      "1133_GTT_DETERMINE_EXCLUSIVITY"(TankID_InOperation := 11, DemandComplete := #GTT_OUT.GTT_DemandsCompleted[11], GTT_Exclusivity := #GTT_Exclusivity)
   END_RUNG
   RUNG wire#powerrail
      { S7_Templates := "SrcType := Int" } EQ_Contact(in1 := #GTT_Exclusivity.TankID_InOperation, in2 := 11)
   END_RUNG wire#w2
   RUNG wire#w2
      I_Coil( #DNC_5S_GTT.Reset )
   END_RUNG
   // the same network as SCL:
   #_w1 := (NOT #GTT_Exclusivity.Tank_Exclusivity AND #GTT_IN.GTT_Actuate[10] AND NOT #GTT_OUT.GTT_DemandsCompleted[10]) OR (#GTT_Exclusivity.TankID_InOperation = 10);
   #"5P_GTT_TimeSel" := "1135_VALVE_OPEN_CLOSE_TIME_SEL"(EN := #_w1,
                           ValveType := 0,
                           ValveDemand := #GTT_IN.GTT_ValveDemands[10],
                           OpenTime := "1096_ADJUSTABLE_CONSTANTS".BWTInletValveOpen_Time,
                           CloseTime := "1096_ADJUSTABLE_CONSTANTS".BWTInletValveClose_Time,
                           ENO => #_w2);
   #DNC_5P_GTT(EN := #_w2,   // "1604_DEMAND_AND_CHECK"
               DemandIn := #GTT_IN.GTT_ValveDemands[10],
               NO_Type := False,
               NC_Type := True,
               ValveMoveTime := #"5P_GTT_TimeSel",
               ValveOpenStatus := "20_TANKS_IP_DATA".RIO_05.FIRST_TANK.TANK_VENT_A_OPEN,
               ValveClsdStatus := "20_TANKS_IP_DATA".RIO_05.FIRST_TANK.TANK_VENT_A_CLSD,
               DemandOut => "40_TANKS_OP_DATA".RIO_05_VENT_A_5P,
               DemandComplete => #GTT_OUT.GTT_DemandsCompleted[10],
               Alarm => #GTT_OUT.GTT_Alarms[10],
               ENO => #_w3);
   IF #_w3 THEN
       "1133_GTT_DETERMINE_EXCLUSIVITY"(TankID_InOperation := 10,
                               DemandComplete := #GTT_OUT.GTT_DemandsCompleted[10],
                               GTT_Exclusivity := #GTT_Exclusivity);
   END_IF;
   #DNC_5P_GTT.Reset := NOT #_w1;
   #_w4 := (NOT #GTT_Exclusivity.Tank_Exclusivity AND #GTT_IN.GTT_Actuate[11] AND NOT #GTT_OUT.GTT_DemandsCompleted[11]) OR (#GTT_Exclusivity.TankID_InOperation = 11);
   #"5S_GTT_TimeSel" := "1135_VALVE_OPEN_CLOSE_TIME_SEL"(EN := #_w4,
                           ValveType := 0,
                           ValveDemand := #GTT_IN.GTT_ValveDemands[11],
                           OpenTime := "1096_ADJUSTABLE_CONSTANTS".BWTInletValveOpen_Time,
                           CloseTime := "1096_ADJUSTABLE_CONSTANTS".BWTInletValveClose_Time,
                           ENO => #_w5);
   #DNC_5S_GTT(EN := #_w5,   // "1604_DEMAND_AND_CHECK"
               DemandIn := #GTT_IN.GTT_ValveDemands[11],
               NO_Type := False,
               NC_Type := True,
               ValveMoveTime := #"5S_GTT_TimeSel",
               ValveOpenStatus := "20_TANKS_IP_DATA".RIO_05.SECOND_TANK.TANK_VENT_A_OPEN,
               ValveClsdStatus := "20_TANKS_IP_DATA".RIO_05.SECOND_TANK.TANK_VENT_A_CLSD,
               DemandOut => "40_TANKS_OP_DATA".RIO_05_VENT_A_5S,
               DemandComplete => #GTT_OUT.GTT_DemandsCompleted[11],
               Alarm => #GTT_OUT.GTT_Alarms[11],
               ENO => #_w6);
   IF #_w6 THEN
       "1133_GTT_DETERMINE_EXCLUSIVITY"(TankID_InOperation := 11,
                               DemandComplete := #GTT_OUT.GTT_DemandsCompleted[11],
                               GTT_Exclusivity := #GTT_Exclusivity);
   END_IF;
   #DNC_5S_GTT.Reset := NOT #_w4;
END_REGION

REGION Network 7: RIO02 6P, 6S GTT control
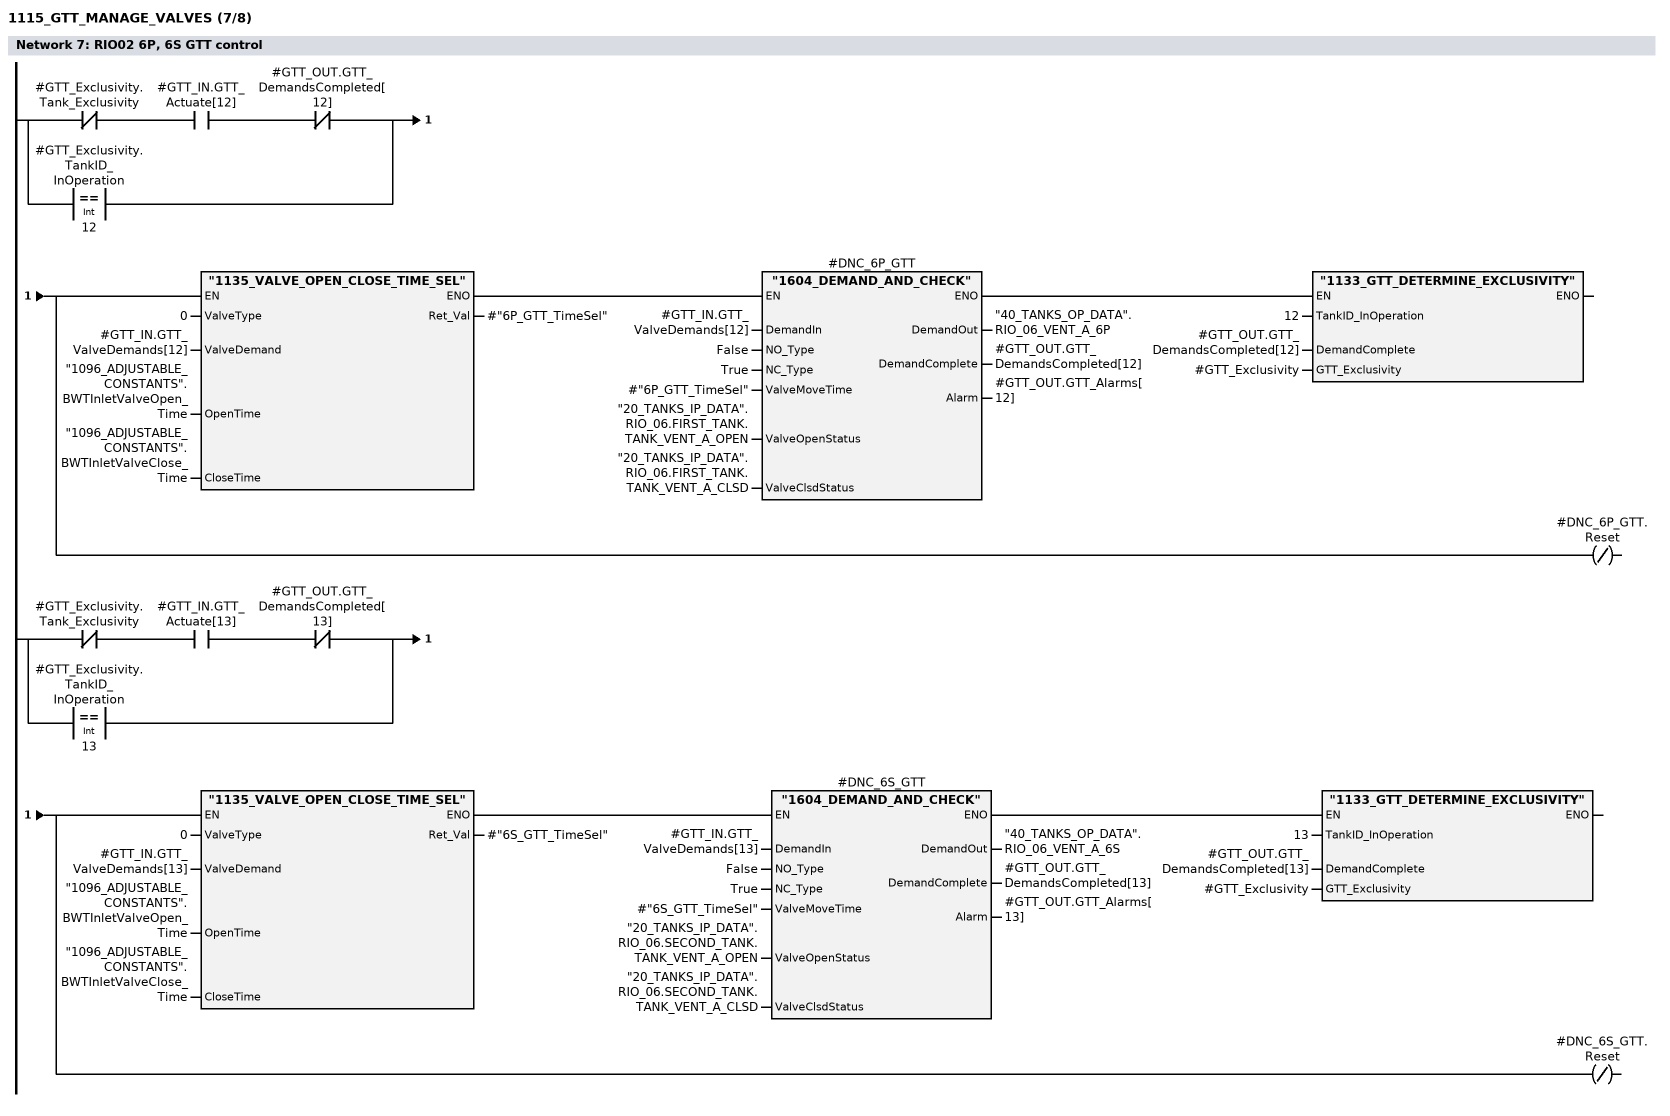
   RUNG wire#powerrail
      I_Contact( #GTT_Exclusivity.Tank_Exclusivity )
      Contact( #GTT_IN.GTT_Actuate[12] )
      I_Contact( #GTT_OUT.GTT_DemandsCompleted[12] )
      wire#w1
      "1135_VALVE_OPEN_CLOSE_TIME_SEL"(ValveType := 0, ValveDemand := #GTT_IN.GTT_ValveDemands[12], OpenTime := "1096_ADJUSTABLE_CONSTANTS".BWTInletValveOpen_Time, CloseTime := "1096_ADJUSTABLE_CONSTANTS".BWTInletValveClose_Time, Ret_Val => #"6P_GTT_TimeSel")
      #DNC_6P_GTT(DemandIn := #GTT_IN.GTT_ValveDemands[12], NO_Type := False, NC_Type := True, ValveMoveTime := #"6P_GTT_TimeSel", ValveOpenStatus := "20_TANKS_IP_DATA".RIO_06.FIRST_TANK.TANK_VENT_A_OPEN, ValveClsdStatus := "20_TANKS_IP_DATA".RIO_06.FIRST_TANK.TANK_VENT_A_CLSD, DemandOut => "40_TANKS_OP_DATA".RIO_06_VENT_A_6P, DemandComplete => #GTT_OUT.GTT_DemandsCompleted[12], Alarm => #GTT_OUT.GTT_Alarms[12])
      "1133_GTT_DETERMINE_EXCLUSIVITY"(TankID_InOperation := 12, DemandComplete := #GTT_OUT.GTT_DemandsCompleted[12], GTT_Exclusivity := #GTT_Exclusivity)
   END_RUNG
   RUNG wire#powerrail
      { S7_Templates := "SrcType := Int" } EQ_Contact(in1 := #GTT_Exclusivity.TankID_InOperation, in2 := 12)
   END_RUNG wire#w1
   RUNG wire#w1
      I_Coil( #DNC_6P_GTT.Reset )
   END_RUNG
   RUNG wire#powerrail
      I_Contact( #GTT_Exclusivity.Tank_Exclusivity )
      Contact( #GTT_IN.GTT_Actuate[13] )
      I_Contact( #GTT_OUT.GTT_DemandsCompleted[13] )
      wire#w2
      "1135_VALVE_OPEN_CLOSE_TIME_SEL"(ValveType := 0, ValveDemand := #GTT_IN.GTT_ValveDemands[13], OpenTime := "1096_ADJUSTABLE_CONSTANTS".BWTInletValveOpen_Time, CloseTime := "1096_ADJUSTABLE_CONSTANTS".BWTInletValveClose_Time, Ret_Val => #"6S_GTT_TimeSel")
      #DNC_6S_GTT(DemandIn := #GTT_IN.GTT_ValveDemands[13], NO_Type := False, NC_Type := True, ValveMoveTime := #"6S_GTT_TimeSel", ValveOpenStatus := "20_TANKS_IP_DATA".RIO_06.SECOND_TANK.TANK_VENT_A_OPEN, ValveClsdStatus := "20_TANKS_IP_DATA".RIO_06.SECOND_TANK.TANK_VENT_A_CLSD, DemandOut => "40_TANKS_OP_DATA".RIO_06_VENT_A_6S, DemandComplete => #GTT_OUT.GTT_DemandsCompleted[13], Alarm => #GTT_OUT.GTT_Alarms[13])
      "1133_GTT_DETERMINE_EXCLUSIVITY"(TankID_InOperation := 13, DemandComplete := #GTT_OUT.GTT_DemandsCompleted[13], GTT_Exclusivity := #GTT_Exclusivity)
   END_RUNG
   RUNG wire#powerrail
      { S7_Templates := "SrcType := Int" } EQ_Contact(in1 := #GTT_Exclusivity.TankID_InOperation, in2 := 13)
   END_RUNG wire#w2
   RUNG wire#w2
      I_Coil( #DNC_6S_GTT.Reset )
   END_RUNG
   // the same network as SCL:
   #_w1 := (NOT #GTT_Exclusivity.Tank_Exclusivity AND #GTT_IN.GTT_Actuate[12] AND NOT #GTT_OUT.GTT_DemandsCompleted[12]) OR (#GTT_Exclusivity.TankID_InOperation = 12);
   #"6P_GTT_TimeSel" := "1135_VALVE_OPEN_CLOSE_TIME_SEL"(EN := #_w1,
                           ValveType := 0,
                           ValveDemand := #GTT_IN.GTT_ValveDemands[12],
                           OpenTime := "1096_ADJUSTABLE_CONSTANTS".BWTInletValveOpen_Time,
                           CloseTime := "1096_ADJUSTABLE_CONSTANTS".BWTInletValveClose_Time,
                           ENO => #_w2);
   #DNC_6P_GTT(EN := #_w2,   // "1604_DEMAND_AND_CHECK"
               DemandIn := #GTT_IN.GTT_ValveDemands[12],
               NO_Type := False,
               NC_Type := True,
               ValveMoveTime := #"6P_GTT_TimeSel",
               ValveOpenStatus := "20_TANKS_IP_DATA".RIO_06.FIRST_TANK.TANK_VENT_A_OPEN,
               ValveClsdStatus := "20_TANKS_IP_DATA".RIO_06.FIRST_TANK.TANK_VENT_A_CLSD,
               DemandOut => "40_TANKS_OP_DATA".RIO_06_VENT_A_6P,
               DemandComplete => #GTT_OUT.GTT_DemandsCompleted[12],
               Alarm => #GTT_OUT.GTT_Alarms[12],
               ENO => #_w3);
   IF #_w3 THEN
       "1133_GTT_DETERMINE_EXCLUSIVITY"(TankID_InOperation := 12,
                               DemandComplete := #GTT_OUT.GTT_DemandsCompleted[12],
                               GTT_Exclusivity := #GTT_Exclusivity);
   END_IF;
   #DNC_6P_GTT.Reset := NOT #_w1;
   #_w4 := (NOT #GTT_Exclusivity.Tank_Exclusivity AND #GTT_IN.GTT_Actuate[13] AND NOT #GTT_OUT.GTT_DemandsCompleted[13]) OR (#GTT_Exclusivity.TankID_InOperation = 13);
   #"6S_GTT_TimeSel" := "1135_VALVE_OPEN_CLOSE_TIME_SEL"(EN := #_w4,
                           ValveType := 0,
                           ValveDemand := #GTT_IN.GTT_ValveDemands[13],
                           OpenTime := "1096_ADJUSTABLE_CONSTANTS".BWTInletValveOpen_Time,
                           CloseTime := "1096_ADJUSTABLE_CONSTANTS".BWTInletValveClose_Time,
                           ENO => #_w5);
   #DNC_6S_GTT(EN := #_w5,   // "1604_DEMAND_AND_CHECK"
               DemandIn := #GTT_IN.GTT_ValveDemands[13],
               NO_Type := False,
               NC_Type := True,
               ValveMoveTime := #"6S_GTT_TimeSel",
               ValveOpenStatus := "20_TANKS_IP_DATA".RIO_06.SECOND_TANK.TANK_VENT_A_OPEN,
               ValveClsdStatus := "20_TANKS_IP_DATA".RIO_06.SECOND_TANK.TANK_VENT_A_CLSD,
               DemandOut => "40_TANKS_OP_DATA".RIO_06_VENT_A_6S,
               DemandComplete => #GTT_OUT.GTT_DemandsCompleted[13],
               Alarm => #GTT_OUT.GTT_Alarms[13],
               ENO => #_w6);
   IF #_w6 THEN
       "1133_GTT_DETERMINE_EXCLUSIVITY"(TankID_InOperation := 13,
                               DemandComplete := #GTT_OUT.GTT_DemandsCompleted[13],
                               GTT_Exclusivity := #GTT_Exclusivity);
   END_IF;
   #DNC_6S_GTT.Reset := NOT #_w4;
END_REGION

REGION Network 8: RIO07 APT GTT control
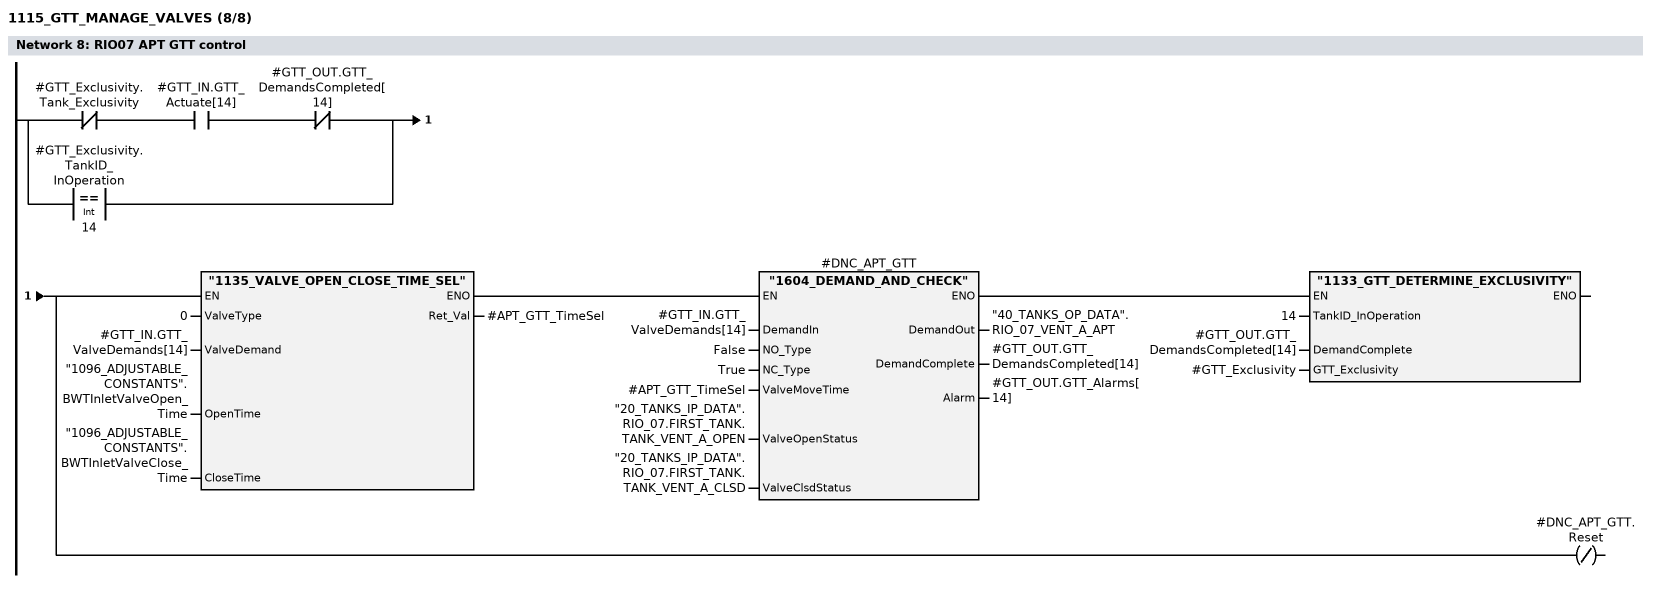
   RUNG wire#powerrail
      I_Contact( #GTT_Exclusivity.Tank_Exclusivity )
      Contact( #GTT_IN.GTT_Actuate[14] )
      I_Contact( #GTT_OUT.GTT_DemandsCompleted[14] )
      wire#w1
      "1135_VALVE_OPEN_CLOSE_TIME_SEL"(ValveType := 0, ValveDemand := #GTT_IN.GTT_ValveDemands[14], OpenTime := "1096_ADJUSTABLE_CONSTANTS".BWTInletValveOpen_Time, CloseTime := "1096_ADJUSTABLE_CONSTANTS".BWTInletValveClose_Time, Ret_Val => #APT_GTT_TimeSel)
      #DNC_APT_GTT(DemandIn := #GTT_IN.GTT_ValveDemands[14], NO_Type := False, NC_Type := True, ValveMoveTime := #APT_GTT_TimeSel, ValveOpenStatus := "20_TANKS_IP_DATA".RIO_07.FIRST_TANK.TANK_VENT_A_OPEN, ValveClsdStatus := "20_TANKS_IP_DATA".RIO_07.FIRST_TANK.TANK_VENT_A_CLSD, DemandOut => "40_TANKS_OP_DATA".RIO_07_VENT_A_APT, DemandComplete => #GTT_OUT.GTT_DemandsCompleted[14], Alarm => #GTT_OUT.GTT_Alarms[14])
      "1133_GTT_DETERMINE_EXCLUSIVITY"(TankID_InOperation := 14, DemandComplete := #GTT_OUT.GTT_DemandsCompleted[14], GTT_Exclusivity := #GTT_Exclusivity)
   END_RUNG
   RUNG wire#powerrail
      { S7_Templates := "SrcType := Int" } EQ_Contact(in1 := #GTT_Exclusivity.TankID_InOperation, in2 := 14)
   END_RUNG wire#w1
   RUNG wire#w1
      I_Coil( #DNC_APT_GTT.Reset )
   END_RUNG
   // the same network as SCL:
   #_w1 := (NOT #GTT_Exclusivity.Tank_Exclusivity AND #GTT_IN.GTT_Actuate[14] AND NOT #GTT_OUT.GTT_DemandsCompleted[14]) OR (#GTT_Exclusivity.TankID_InOperation = 14);
   #APT_GTT_TimeSel := "1135_VALVE_OPEN_CLOSE_TIME_SEL"(EN := #_w1,
                           ValveType := 0,
                           ValveDemand := #GTT_IN.GTT_ValveDemands[14],
                           OpenTime := "1096_ADJUSTABLE_CONSTANTS".BWTInletValveOpen_Time,
                           CloseTime := "1096_ADJUSTABLE_CONSTANTS".BWTInletValveClose_Time,
                           ENO => #_w2);
   #DNC_APT_GTT(EN := #_w2,   // "1604_DEMAND_AND_CHECK"
                DemandIn := #GTT_IN.GTT_ValveDemands[14],
                NO_Type := False,
                NC_Type := True,
                ValveMoveTime := #APT_GTT_TimeSel,
                ValveOpenStatus := "20_TANKS_IP_DATA".RIO_07.FIRST_TANK.TANK_VENT_A_OPEN,
                ValveClsdStatus := "20_TANKS_IP_DATA".RIO_07.FIRST_TANK.TANK_VENT_A_CLSD,
                DemandOut => "40_TANKS_OP_DATA".RIO_07_VENT_A_APT,
                DemandComplete => #GTT_OUT.GTT_DemandsCompleted[14],
                Alarm => #GTT_OUT.GTT_Alarms[14],
                ENO => #_w3);
   IF #_w3 THEN
       "1133_GTT_DETERMINE_EXCLUSIVITY"(TankID_InOperation := 14,
                               DemandComplete := #GTT_OUT.GTT_DemandsCompleted[14],
                               GTT_Exclusivity := #GTT_Exclusivity);
   END_IF;
   #DNC_APT_GTT.Reset := NOT #_w1;
END_REGION
END_FUNCTION_BLOCK

FUNCTION_BLOCK "1120_PVV_MANAGE_VALVES"   // FB1120, LAD
{ S7_Optimized_Access := 'TRUE' }
VERSION : 0.1
// Manage the Vent A and Vent B valves based on the provided data.
// "Actuate" enables the actuation of the valves in question (grouped A and B).
// "ValveDemands" signifies whether the valve should be actuating (Openning as NC valve) or releasing (Closing as NC valve).
// 
// This function puts out two sets of data:
// "DemandsCompleted" which indicates whether the demand is complete.
// "Alarms" indicated if an alarm has been triggered (e.g. a timeout in the Demand And Check.
// 
// The timeout for Demand and Check is automatically selected based on the demand and valve type.
   VAR_INPUT
      PVVX_IN : "VALVE_PVVX_IN";
   END_VAR
   VAR_OUTPUT
      PVVX_OUT : "VALVE_PVVX_OUT";
   END_VAR
   VAR
      DNC_FPT_VENTA : "1604_DEMAND_AND_CHECK";
      DNC_FPT_VENTB : "1604_DEMAND_AND_CHECK";
      DNC_1P_VENTA : "1604_DEMAND_AND_CHECK";
      DNC_1P_VENTB : "1604_DEMAND_AND_CHECK";
      DNC_1S_VENTA : "1604_DEMAND_AND_CHECK";
      DNC_1S_VENTB : "1604_DEMAND_AND_CHECK";
      DNC_2P_VENTA : "1604_DEMAND_AND_CHECK";
      DNC_2P_VENTB : "1604_DEMAND_AND_CHECK";
      DNC_2S_VENTA : "1604_DEMAND_AND_CHECK";
      DNC_2S_VENTB : "1604_DEMAND_AND_CHECK";
      DNC_3P_VENTA : "1604_DEMAND_AND_CHECK";
      DNC_3P_VENTB : "1604_DEMAND_AND_CHECK";
      DNC_3S_VENTA : "1604_DEMAND_AND_CHECK";
      DNC_3S_VENTB : "1604_DEMAND_AND_CHECK";
      DNC_4P_VENTA : "1604_DEMAND_AND_CHECK";
      DNC_4P_VENTB : "1604_DEMAND_AND_CHECK";
      DNC_4S_VENTA : "1604_DEMAND_AND_CHECK";
      DNC_4S_VENTB : "1604_DEMAND_AND_CHECK";
      DNC_5P_VENTA : "1604_DEMAND_AND_CHECK";
      DNC_5P_VENTB : "1604_DEMAND_AND_CHECK";
      DNC_5S_VENTA : "1604_DEMAND_AND_CHECK";
      DNC_5S_VENTB : "1604_DEMAND_AND_CHECK";
      DNC_6P_VENTA : "1604_DEMAND_AND_CHECK";
      DNC_6P_VENTB : "1604_DEMAND_AND_CHECK";
      DNC_6S_VENTA : "1604_DEMAND_AND_CHECK";
      DNC_6S_VENTB : "1604_DEMAND_AND_CHECK";
      DNC_APT_VENTA : "1604_DEMAND_AND_CHECK";
      DNC_APT_VENTB : "1604_DEMAND_AND_CHECK";
   END_VAR
   VAR_TEMP
      FPT_VentA_TimeSel : Time;
      FPT_VentB_TimeSel : Time;
      "1P_VentA_TimeSel" : Time;
      "1P_VentB_TimeSel" : Time;
      "1S_VentA_TimeSel" : Time;
      "1S_VentB_TimeSel" : Time;
      "2P_VentA_TimeSel" : Time;
      "2P_VentB_TimeSel" : Time;
      "2S_VentA_TimeSel" : Time;
      "2S_VentB_TimeSel" : Time;
      "3P_VentA_TimeSel" : Time;
      "3P_VentB_TimeSel" : Time;
      "3S_VentA_TimeSel" : Time;
      "3S_VentB_TimeSel" : Time;
      "4P_VentA_TimeSel" : Time;
      "4P_VentB_TimeSel" : Time;
      "4S_VentA_TimeSel" : Time;
      "4S_VentB_TimeSel" : Time;
      "5P_VentA_TimeSel" : Time;
      "5P_VentB_TimeSel" : Time;
      "5S_VentA_TimeSel" : Time;
      "5S_VentB_TimeSel" : Time;
      "6P_VentA_TimeSel" : Time;
      "6P_VentB_TimeSel" : Time;
      "6S_VentA_TimeSel" : Time;
      "6S_VentB_TimeSel" : Time;
      APT_VentA_TimeSel : Time;
      APT_VentB_TimeSel : Time;
   END_VAR
   VAR CONSTANT
      TimerResetHold : LTime := LT#30s;
   END_VAR
   VAR_TEMP   // added for the SCL form of the ladder/FBD networks
      _w1 : Bool;
      _w2 : Bool;
      _w3 : Bool;
      _w4 : Bool;
      _w5 : Bool;
      _w6 : Bool;
      _w7 : Bool;
      _w8 : Bool;
      _w9 : Bool;
   END_VAR
BEGIN

REGION Network 1: Reset all timers if they are not in actuation mode.
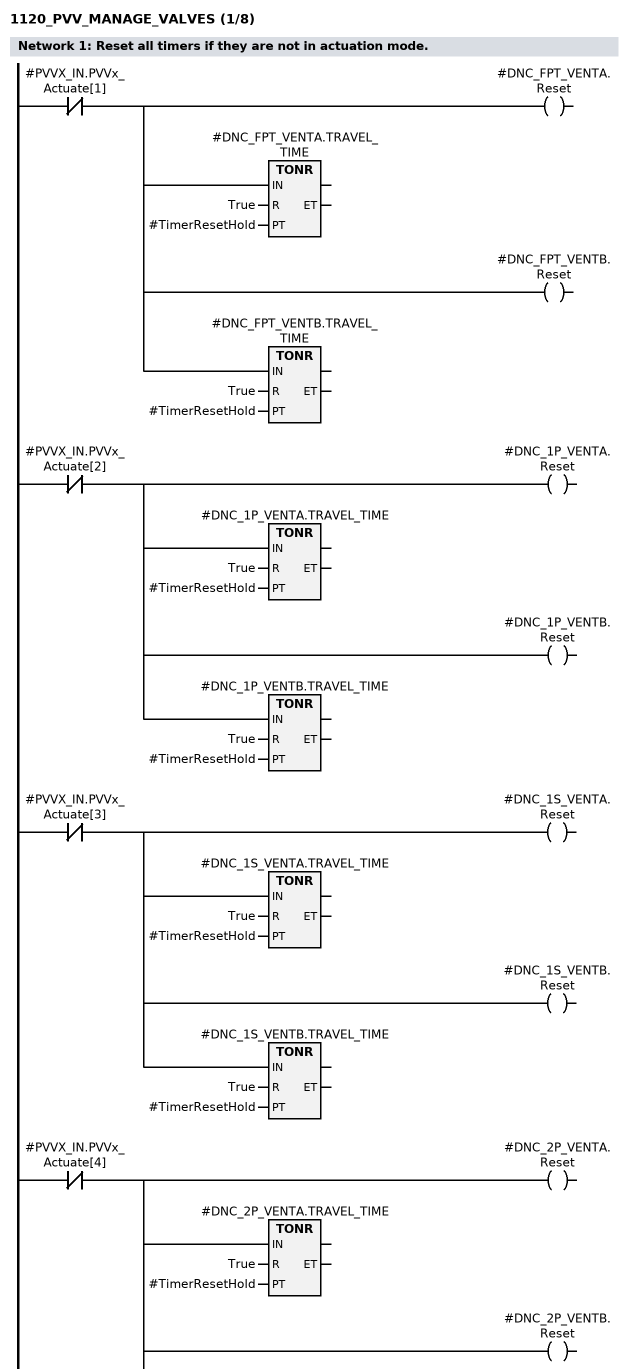
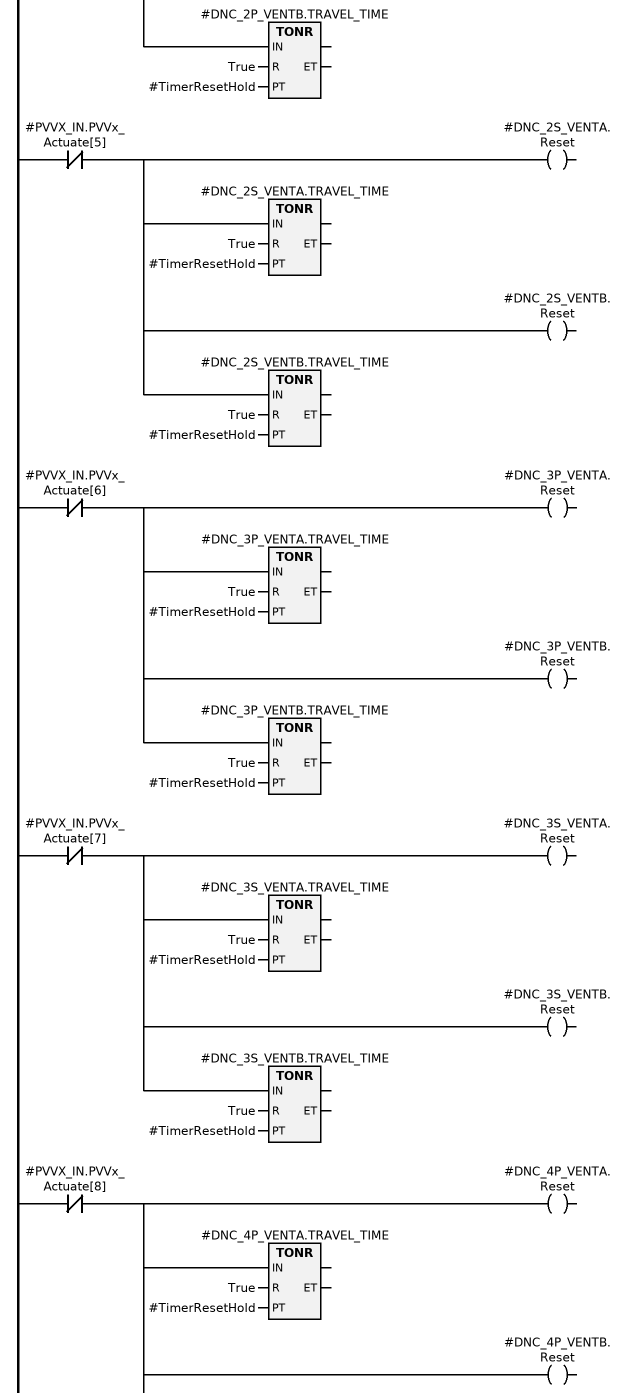
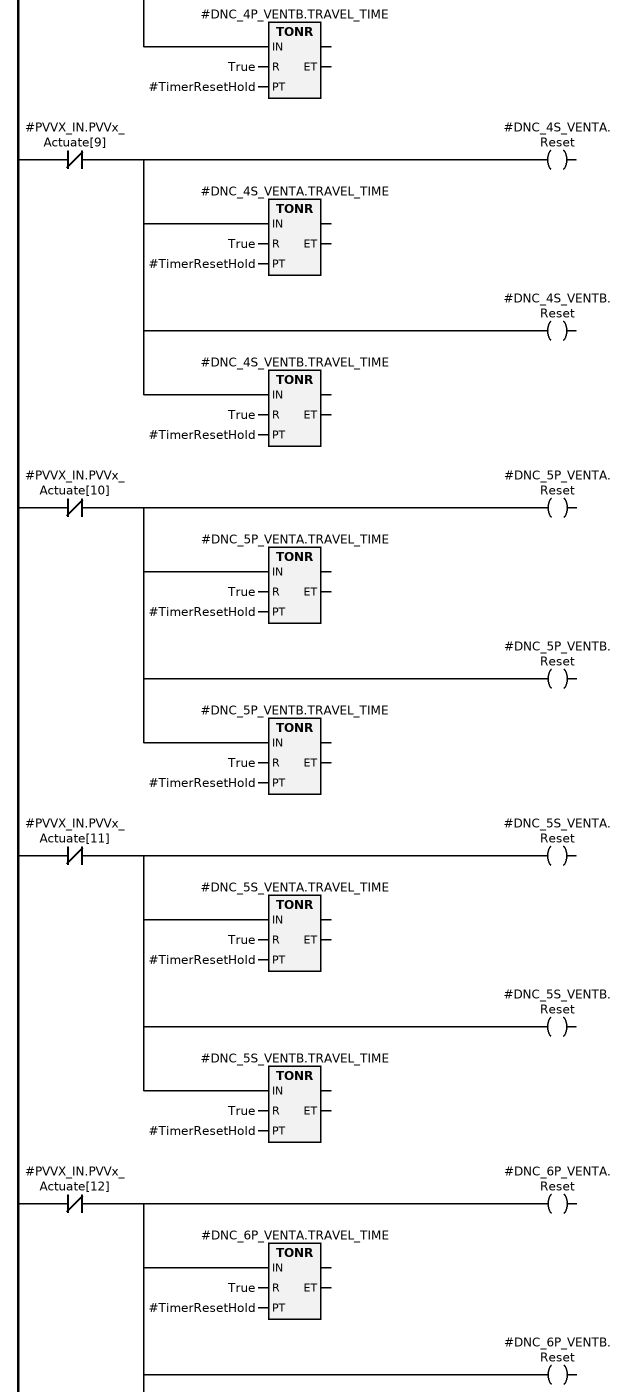
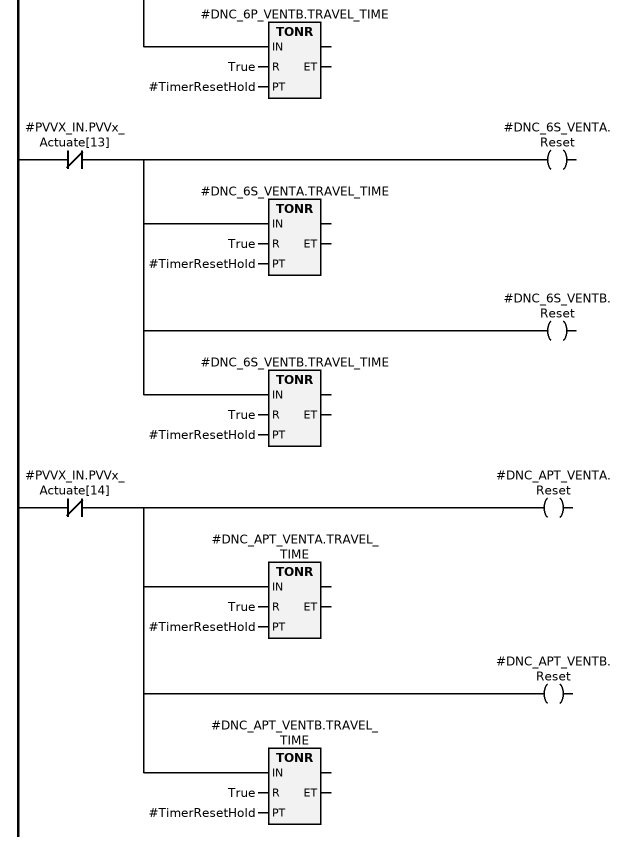
   #DNC_FPT_VENTA.Reset := NOT #PVVX_IN.PVVx_Actuate[1];
   #DNC_FPT_VENTA.TRAVEL_TIME.TONR(IN := NOT #PVVX_IN.PVVx_Actuate[1], R := True, PT := #TimerResetHold);
   #DNC_FPT_VENTB.Reset := NOT #PVVX_IN.PVVx_Actuate[1];
   #DNC_FPT_VENTB.TRAVEL_TIME.TONR(IN := NOT #PVVX_IN.PVVx_Actuate[1], R := True, PT := #TimerResetHold);
   #DNC_1P_VENTA.Reset := NOT #PVVX_IN.PVVx_Actuate[2];
   #DNC_1P_VENTA.TRAVEL_TIME.TONR(IN := NOT #PVVX_IN.PVVx_Actuate[2], R := True, PT := #TimerResetHold);
   #DNC_1P_VENTB.Reset := NOT #PVVX_IN.PVVx_Actuate[2];
   #DNC_1P_VENTB.TRAVEL_TIME.TONR(IN := NOT #PVVX_IN.PVVx_Actuate[2], R := True, PT := #TimerResetHold);
   #DNC_1S_VENTA.Reset := NOT #PVVX_IN.PVVx_Actuate[3];
   #DNC_1S_VENTA.TRAVEL_TIME.TONR(IN := NOT #PVVX_IN.PVVx_Actuate[3], R := True, PT := #TimerResetHold);
   #DNC_1S_VENTB.Reset := NOT #PVVX_IN.PVVx_Actuate[3];
   #DNC_1S_VENTB.TRAVEL_TIME.TONR(IN := NOT #PVVX_IN.PVVx_Actuate[3], R := True, PT := #TimerResetHold);
   #DNC_2P_VENTA.Reset := NOT #PVVX_IN.PVVx_Actuate[4];
   #DNC_2P_VENTA.TRAVEL_TIME.TONR(IN := NOT #PVVX_IN.PVVx_Actuate[4], R := True, PT := #TimerResetHold);
   #DNC_2P_VENTB.Reset := NOT #PVVX_IN.PVVx_Actuate[4];
   #DNC_2P_VENTB.TRAVEL_TIME.TONR(IN := NOT #PVVX_IN.PVVx_Actuate[4], R := True, PT := #TimerResetHold);
   #DNC_2S_VENTA.Reset := NOT #PVVX_IN.PVVx_Actuate[5];
   #DNC_2S_VENTA.TRAVEL_TIME.TONR(IN := NOT #PVVX_IN.PVVx_Actuate[5], R := True, PT := #TimerResetHold);
   #DNC_2S_VENTB.Reset := NOT #PVVX_IN.PVVx_Actuate[5];
   #DNC_2S_VENTB.TRAVEL_TIME.TONR(IN := NOT #PVVX_IN.PVVx_Actuate[5], R := True, PT := #TimerResetHold);
   #DNC_3P_VENTA.Reset := NOT #PVVX_IN.PVVx_Actuate[6];
   #DNC_3P_VENTA.TRAVEL_TIME.TONR(IN := NOT #PVVX_IN.PVVx_Actuate[6], R := True, PT := #TimerResetHold);
   #DNC_3P_VENTB.Reset := NOT #PVVX_IN.PVVx_Actuate[6];
   #DNC_3P_VENTB.TRAVEL_TIME.TONR(IN := NOT #PVVX_IN.PVVx_Actuate[6], R := True, PT := #TimerResetHold);
   #DNC_3S_VENTA.Reset := NOT #PVVX_IN.PVVx_Actuate[7];
   #DNC_3S_VENTA.TRAVEL_TIME.TONR(IN := NOT #PVVX_IN.PVVx_Actuate[7], R := True, PT := #TimerResetHold);
   #DNC_3S_VENTB.Reset := NOT #PVVX_IN.PVVx_Actuate[7];
   #DNC_3S_VENTB.TRAVEL_TIME.TONR(IN := NOT #PVVX_IN.PVVx_Actuate[7], R := True, PT := #TimerResetHold);
   #DNC_4P_VENTA.Reset := NOT #PVVX_IN.PVVx_Actuate[8];
   #DNC_4P_VENTA.TRAVEL_TIME.TONR(IN := NOT #PVVX_IN.PVVx_Actuate[8], R := True, PT := #TimerResetHold);
   #DNC_4P_VENTB.Reset := NOT #PVVX_IN.PVVx_Actuate[8];
   #DNC_4P_VENTB.TRAVEL_TIME.TONR(IN := NOT #PVVX_IN.PVVx_Actuate[8], R := True, PT := #TimerResetHold);
   #DNC_4S_VENTA.Reset := NOT #PVVX_IN.PVVx_Actuate[9];
   #DNC_4S_VENTA.TRAVEL_TIME.TONR(IN := NOT #PVVX_IN.PVVx_Actuate[9], R := True, PT := #TimerResetHold);
   #DNC_4S_VENTB.Reset := NOT #PVVX_IN.PVVx_Actuate[9];
   #DNC_4S_VENTB.TRAVEL_TIME.TONR(IN := NOT #PVVX_IN.PVVx_Actuate[9], R := True, PT := #TimerResetHold);
   #DNC_5P_VENTA.Reset := NOT #PVVX_IN.PVVx_Actuate[10];
   #DNC_5P_VENTA.TRAVEL_TIME.TONR(IN := NOT #PVVX_IN.PVVx_Actuate[10], R := True, PT := #TimerResetHold);
   #DNC_5P_VENTB.Reset := NOT #PVVX_IN.PVVx_Actuate[10];
   #DNC_5P_VENTB.TRAVEL_TIME.TONR(IN := NOT #PVVX_IN.PVVx_Actuate[10], R := True, PT := #TimerResetHold);
   #DNC_5S_VENTA.Reset := NOT #PVVX_IN.PVVx_Actuate[11];
   #DNC_5S_VENTA.TRAVEL_TIME.TONR(IN := NOT #PVVX_IN.PVVx_Actuate[11], R := True, PT := #TimerResetHold);
   #DNC_5S_VENTB.Reset := NOT #PVVX_IN.PVVx_Actuate[11];
   #DNC_5S_VENTB.TRAVEL_TIME.TONR(IN := NOT #PVVX_IN.PVVx_Actuate[11], R := True, PT := #TimerResetHold);
   #DNC_6P_VENTA.Reset := NOT #PVVX_IN.PVVx_Actuate[12];
   #DNC_6P_VENTA.TRAVEL_TIME.TONR(IN := NOT #PVVX_IN.PVVx_Actuate[12], R := True, PT := #TimerResetHold);
   #DNC_6P_VENTB.Reset := NOT #PVVX_IN.PVVx_Actuate[12];
   #DNC_6P_VENTB.TRAVEL_TIME.TONR(IN := NOT #PVVX_IN.PVVx_Actuate[12], R := True, PT := #TimerResetHold);
   #DNC_6S_VENTA.Reset := NOT #PVVX_IN.PVVx_Actuate[13];
   #DNC_6S_VENTA.TRAVEL_TIME.TONR(IN := NOT #PVVX_IN.PVVx_Actuate[13], R := True, PT := #TimerResetHold);
   #DNC_6S_VENTB.Reset := NOT #PVVX_IN.PVVx_Actuate[13];
   #DNC_6S_VENTB.TRAVEL_TIME.TONR(IN := NOT #PVVX_IN.PVVx_Actuate[13], R := True, PT := #TimerResetHold);
   #DNC_APT_VENTA.Reset := NOT #PVVX_IN.PVVx_Actuate[14];
   #DNC_APT_VENTA.TRAVEL_TIME.TONR(IN := NOT #PVVX_IN.PVVx_Actuate[14], R := True, PT := #TimerResetHold);
   #DNC_APT_VENTB.Reset := NOT #PVVX_IN.PVVx_Actuate[14];
   #DNC_APT_VENTB.TRAVEL_TIME.TONR(IN := NOT #PVVX_IN.PVVx_Actuate[14], R := True, PT := #TimerResetHold);
END_REGION

REGION Network 2: RIO01 FPT, 1P, 1S Vent A and Vent B control